FUNCTION "LOWERCASE" : String[254]   // FC273, SCL
TITLE = LOWERCASE
{ S7_Optimized_Access := 'FALSE' }
AUTHOR : hugo
FAMILY : STRINGS
NAME : LOWCASE
VERSION : 1.3
// lowercase returns str while all letters A..Z and Ä.Ö,Ü are converted to lowercase.
//  
// uses: SETUP [DB1]
//       TO_LOWER [FC282]
   VAR_INPUT
      str : String[254];
      _str AT str : Struct
         length : Byte;
         act_length : Byte;
         str : Array[1..254] of Byte;
      END_STRUCT;
   END_VAR
   VAR_TEMP
      tLOWERCASE : String[254];
      _LOWERCASE AT tLOWERCASE : Struct
         length : Byte;
         act_length : Byte;
         str : Array[1..254] of Byte;
      END_STRUCT;
      PT : Int;   // PT : POINTER TO BYTE;
      pos : Int;
      l : Int;
   END_VAR
BEGIN


   #PT := 1;                                    //ADR(LOWERCASE);
   #tLOWERCASE := #str;
   #l := BYTE_TO_INT(#_LOWERCASE.act_length);    //LEN(str);
   FOR #pos := 1 TO #l DO
       #_LOWERCASE.str[#PT] := "TO_LOWER"(#_LOWERCASE.str[#PT]);
       #PT := #PT + 1;
   END_FOR;

   #LOWERCASE := #tLOWERCASE;

   (* revision histroy
   hm  6. oct. 2006    rev 1.0
       original release

   hm  4. feb. 2008    rev 1.1
       improved performance
       added Ä.Ö,Ü

   hm  6. mar. 2008    rev 1.2
       added support for exteded Ascii

   hm  29. mar. 2008   rev 1.3
       changed STRING to STRING(STRING_LENGTH)
   *)
END_FUNCTION

FUNCTION "MIRROR" : String[254]   // FC274, SCL
TITLE = MIRROR
{ S7_Optimized_Access := 'FALSE' }
AUTHOR : hugo
FAMILY : STRINGS
NAME : MIRROR
VERSION : 1.1
// this function reverses an input string.
   VAR_INPUT
      str : String[254];
      _str AT str : Struct
         length : Byte;
         act_length : Byte;
         str : Array[1..254] of Byte;
      END_STRUCT;
   END_VAR
   VAR_TEMP
      tmirror : String[254];
      _mirror AT tmirror : Struct
         length : Byte;
         act_length : Byte;
         str : Array[1..254] of Byte;
      END_STRUCT;
      pi : Int;   // pi : POINTER TO ARRAY[1..255] OF BYTE;
      po : Int;   // po : POINTER TO BYTE;
      lx : Int;
      i : Int;
   END_VAR
BEGIN


   #tmirror := #str;

   #pi := 1;    //ADR(str);
   #po := 1;    //ADR(mirror);
   #lx := BYTE_TO_INT(#_str.act_length); //LEN(str);
   FOR #i := #lx TO 1 BY - 1 DO
       #_mirror.str[#po] := #_str.str[#i];
       #po := #po + 1;
   END_FOR;
   (* close output string *)
   //po^:= 0;
   #MIRROR:= #tmirror;


   (* revision histroy
   hm  4. feb. 2008    rev 1.0
       original release

   hm  29. mar. 2008   rev 1.1
       changed STRING to STRING(STRING_LENGTH)
   *)
END_FUNCTION

FUNCTION "MONTH_TO_STRING" : String[254]   // FC275, SCL
TITLE = MONTH_TO_STRING
{ S7_Optimized_Access := 'FALSE' }
AUTHOR : hugo
FAMILY : STRINGS
NAME : MONTHSTR
VERSION : 1.1
// MONTH_TO_STRING converts an Integer 1..12 into a String with the Names of the corresponding Month.
// the decoding is according to the language setup in global vars
// 
// uses: LANGUAGE [DB4]
   VAR_INPUT
      MTH : Int;
      LANG : Int;
      LX : Int;
   END_VAR
   VAR_TEMP
      ly : Int;
   END_VAR
BEGIN


   #MONTH_TO_STRING := ' ';

   IF #LANG = 0 THEN #ly := "LANGUAGE".DEFAULT; ELSE #ly := MIN(IN1:=#LANG, IN2:="LANGUAGE".LMAX); END_IF;
   IF #MTH < 1 OR #MTH > 12 THEN
       RETURN;
   ELSIF #LX = 0 THEN
       #MONTH_TO_STRING := "LANGUAGE".MONTHS[#ly, #MTH];
   ELSIF #LX = 3 THEN
       #MONTH_TO_STRING := "LANGUAGE".MONTHS3[#ly, #MTH];
   END_IF;


   (* revisison history

   hm  21. sep. 2008   rev 1.0
       original version

   hm  19. oct. 2008   rev 1.1
       changed language setup constants
   *)
END_FUNCTION

FUNCTION "OCT_TO_BYTE" : Byte   // FC276, SCL
TITLE = OCT_TO_BYTE
{ S7_Optimized_Access := 'FALSE' }
AUTHOR : hugo
FAMILY : STRINGS
NAME : OCT2BY
VERSION : 1.1
// OCT_TO_BYTE converts a octagonal string into a byte.
   VAR_INPUT
      OCT : String[254];
      _OCT AT OCT : Struct
         length : Byte;
         act_length : Byte;
         str : Array[1..10] of Byte;
      END_STRUCT;
   END_VAR
   VAR_TEMP
      pt : Int;   // pt : POINTER TO BYTE;
      i : Int;
      X : Byte;
      stop : Int;
   END_VAR
BEGIN


   #pt := 1;    //ADR(oct);
   #stop := BYTE_TO_INT(#_OCT.act_length);    //LEN(oct);
   FOR #i := 1 TO #stop DO
       (* read the first character and subtract 48 to get value in decimal 0 = 48 *)
       #X := #_OCT.str[#pt];
       (* calculate the value of the digit *)
       IF BYTE_TO_INT(#X) > 47 AND BYTE_TO_INT(#X) < 56 THEN
           #OCT_TO_BYTE := INT_TO_BYTE(BYTE_TO_INT(SHL(IN:=#OCT_TO_BYTE,N:=3)) + BYTE_TO_INT(#X) - 48);
       END_IF;
       #pt := #pt + 1;
   END_FOR;



   (* revision histroy
   hm  18. jun. 2008   rev 1.0
       original release

   hm  20. sep. 2008   rev 1.1
       changed length of input string from 20 to 10

   *)
END_FUNCTION

FUNCTION "OCT_TO_DWORD" : DWord   // FC277, SCL
TITLE = OCT_TO_DWORD
{ S7_Optimized_Access := 'FALSE' }
AUTHOR : hugo
FAMILY : STRINGS
NAME : OCT2DW
VERSION : 1.0
// OCT_TO_DWORD converts a octagonal string into a dword.
   VAR_INPUT
      OCT : String[254];
      _OCT AT OCT : Struct
         length : Byte;
         act_length : Byte;
         str : Array[1..20] of Byte;
      END_STRUCT;
   END_VAR
   VAR_TEMP
      pt : Int;   // pt : POINTER TO BYTE;
      i : Int;
      X : Byte;
      stop : Int;
   END_VAR
BEGIN


   #pt := 1;    //ADR(oct);
   #stop := BYTE_TO_INT(#_OCT.act_length);   //LEN(oct);
   FOR #i := 1 TO #stop DO
       (* read the first character and subtract 48 to get value in decimal 0 = 48 *)
       #X := #_OCT.str[#pt];
       (* calculate the value of the digit *)
       IF BYTE_TO_INT(#X) > 47 AND BYTE_TO_INT(#X) < 56 THEN
           #OCT_TO_DWORD := DINT_TO_DWORD(DWORD_TO_DINT(SHL(IN:=#OCT_TO_DWORD,N:=3)) + BYTE_TO_INT(#X) - 48);
       END_IF;
       #pt := #pt + 1;
   END_FOR;




   (* revision histroy
   hm  18. jun. 2008   rev 1.0
       original release


   *)
END_FUNCTION

FUNCTION "REAL_TO_STRF" : String[254]   // FC278, SCL
TITLE = REAL_TO_STRF
{ S7_Optimized_Access := 'FALSE' }
AUTHOR : oscat
FAMILY : STRINGS
NAME : REALSTR
VERSION : 1.7
// Real_to_strF converts a Real to a fixed length String.
// the string will be filles with zeroes to achieve the fixed length after the dot.
// 
// uses: DI_STRNG [FC5]
//       CONCAT [FC2]
//       EXP10 [FC77]
//       DELETE [FC4]
//       INSERT [FC17]
   VAR_INPUT
      IN : Real;
      N : Int;
   END_VAR
   VAR_TEMP
      tN : Int;
      O : Real;
      i : Int;
      str : String[20];
      _str AT str : Struct
         length : Byte;
         act_length : Byte;
         str : Array[1..20] of Byte;
      END_STRUCT;
      tStr : String[20];
   END_VAR
BEGIN


   (* Initialisierung der temporären Strings *)
   #str := '';
   #tStr := '';
   (* round the input to N digits and convert to string *)
   (* LIMIT N to 0 .. 7 *)
   #tN := LIMIT(MN:=0,IN:=#N,MX:=7);
   (* round the input to N digits and convert to string *)
   #O := ABS(#IN) * "EXP10"(#tN);
   #str := S_CONV(REAL_TO_DINT(#O));
   (* Vorzeichen löschen *)
   #tStr := DELETE(IN:=#str, L:=1, P:=1); 
   #str BLKMOV #tStr;
   (* add zeroes in front to make sure sting is at least 8 digits long *)
   FOR #i := BYTE_TO_INT(#_str.act_length) TO #tN DO 
       #tStr := CONCAT(IN1:='0', IN2:=#str);
       #str BLKMOV #tStr; 
   END_FOR;
   (* add a dot if n > 0 *)
   IF #IN <> 0 THEN 
       #tStr := INSERT(IN1:=#str, IN2:='.', P:=BYTE_TO_INT(#_str.act_length) - #tN); 
   END_IF;
   #str BLKMOV #tStr;
   (* add a minus sign if in is negative *)
   IF #IN < 0 THEN 
       #str := CONCAT(IN1:='-', IN2:=#tStr); 
   END_IF;

   #REAL_TO_STRF := #str;


   (* revision history
   hm  26 jan 2007 rev 1.0
       original version

   hm  20. nov. 2007   rev 1.1
       when N=0 ther will be no dot at the end of the string.

   hm  15. dec. 2007   rev 1.2
       changed code for better performance

   hm  4. mar. 2008    rev 1.3
       result is now rounded instead of trunc

   hm  20. mar. 2008   rev 1.4
       changed trunc to real_to_dint because trunc was generating wrong values on wago 842

   hm  29. mar. 2008   rev 1.5
       changed STRING to STRING(20)

   hm  4. apr. 2008    rev 1.6
       added variable O to avoid an error uner CoDeSys SP PLCWinNT V2.4

   hm  27. feb. 2009   rev 1.7
       added a missing zero for IN < 1

   *)
END_FUNCTION

FUNCTION "REPLACE_ALL" : String[254]   // FC279, SCL
TITLE = REPLACE_ALL
{ S7_Optimized_Access := 'FALSE' }
AUTHOR : hugo
FAMILY : STRINGS
NAME : REPLALL
VERSION : 1.1
// the function findP searches a string str for the occurence of src beginning at the position pos.
// 
// uses: LEN [FC21]
//       FINDP [FC248]
//       EQ_STRNG [FC10] 
//       MID [FC26] 
//       REPLACE [FC31]
   VAR_INPUT
      str : String[254];
      src : String[254];
      rep : String[254];
   END_VAR
   VAR_TEMP
      tstr : String[254];
      tsrc : String[254];
      trep : String[254];
      tREPLACE_ALL : String[254];
      pos : Int;
      lp : Int;
      lx : Int;
   END_VAR
BEGIN


   #tstr := #str;
   #tsrc := #src;
   #trep := #rep;

   #tREPLACE_ALL := #str;
   #lx := LEN(#tsrc);
   #lp := LEN(#trep);
   #pos := "FINDP"(str:=#tREPLACE_ALL,src:=#tsrc,pos:=1);
   WHILE #pos > 0 DO
       #tREPLACE_ALL := REPLACE(IN1:=#tREPLACE_ALL,IN2:=#trep,L:=#lx,P:=#pos);
       #pos := "FINDP"(str:=#tREPLACE_ALL,src:=#tsrc,pos:=#pos + #lp);
   END_WHILE;

   #REPLACE_ALL := #tREPLACE_ALL;

   (* revision histroy
   hm  4. feb. 2008    rev 1.0
       original release

   hm  29. mar. 2008   rev 1.1
       changed STRING to STRING(STRING_LENGTH)
   *)
END_FUNCTION

FUNCTION "REPLACE_CHARS" : String[254]   // FC280, SCL
TITLE = REPLACE_CHARS
{ S7_Optimized_Access := 'FALSE' }
AUTHOR : hugo
FAMILY : STRINGS
NAME : REPLCHR
VERSION : 1.0
// REPLACE_CHARS erstezt alle character die im string src aufgeführt sind mit dem an der selben stelle im string rep gelisteten character.
// 
// uses: TEMP [DB7]
//       LEN [FC21]
//       LEFT [FC20]
//       MID [FC26]
//       FIND [FC11]
//       REPLACE [FC31]
   VAR_INPUT
      STR : String[254];
      SRC : String[254];
      REP : String[254];
   END_VAR
   VAR_TEMP
      "a" : Int;
      "b" : Int;
      c : String[1];
      stp : Int;
   END_VAR
BEGIN


   "TEMP".STR1 := #STR;
   "TEMP".STR2 := #SRC;
   "TEMP".STR3 := #REP;

   "TEMP".TEMP := #STR;
   (* make sure rep and src are of same length and length is > 0 *)
   #"a" := LEN("TEMP".STR1);
   #"b" := LEN("TEMP".STR3);
   IF #"a" < #"b" THEN
       "TEMP".STR3 := LEFT(IN:="TEMP".STR3, L:=#"a");
   ELSIF #"b" < #"a" THEN
       "TEMP".STR2 := LEFT(IN:="TEMP".STR2, L:=#"b");
   END_IF;

   (* search the string and replace if necessary *)
   #stp := LEN("TEMP".STR1);
   FOR #"a" := 1 TO #stp DO
       #c := MID(IN:="TEMP".TEMP, L:=1, P:=#"a");
       #"b" := FIND(IN1:="TEMP".STR2, IN2:=#c);
       IF #"b" > 0 THEN
           "TEMP".TEMP := REPLACE(IN1:="TEMP".TEMP, IN2:=MID(IN:="TEMP".STR3, L:=1, P:=#"b"), L:=1, P:=#"a");
       END_IF;
   END_FOR;

   #REPLACE_CHARS := "TEMP".TEMP;

   (* revision history
   hm      14. may. 2008   rev 1.0
       original version

   *)
END_FUNCTION

FUNCTION "REPLACE_UML" : String[254]   // FC281, SCL
TITLE = REPLACE_UML
{ S7_Optimized_Access := 'FALSE' }
AUTHOR : kurt
FAMILY : STRINGS
NAME : REPLUML
VERSION : 1.1
// REPLACE_UML replaces all occurences of Ä,Ö,Ü and ä,ö,ü,ß with Ae, ae, Oe, oe, Ue, ue and ss.
// 
// uses: TO_UML [FC283]
//       CHR_TO_STRING [FC227]
   VAR_INPUT
      str : String[254];
      _str AT str : Struct
         length : Byte;
         act_length : Byte;
         str : Array[1..254] of Byte;
      END_STRUCT;
   END_VAR
   VAR_TEMP
      tREPLACE_UML : String[254];
      _REPLACE_UML AT tREPLACE_UML : Struct
         length : Byte;
         act_length : Byte;
         str : Array[1..254] of Byte;
      END_STRUCT;
      l : Int;
      pt : Int;   // pt : POINTER TO BYTE;
      pto : Int;   // pto : POINTER TO BYTE;
      ptm : Int;   // ptm : POINTER TO BYTE;
      pt1 : Int;   // pt1, pt2 : POINTER TO BYTE;
      pt2 : Int;   // pt1, pt2 : POINTER TO BYTE;
      su : String[2];
      _su AT su : Struct
         length : Byte;
         act_length : Byte;
         str : Array[1..2] of Byte;
      END_STRUCT;
      pos : Int;
   END_VAR
BEGIN


   #tREPLACE_UML := #str;

   #pt := 1;    //ADR(str);
   #pto := 1;   //ADR(REPLACE_UML);
   #ptm := #pto; // + INT_TO_DWORD(string_length);
   #pt1 := 1;   //ADR(su);
   #pt2 := #pt1 + 1;
   #l := BYTE_TO_INT(#_str.act_length);   //LEN(str);
   WHILE #pos < #l AND #pos < BYTE_TO_INT(#_str.act_length) DO
       IF BYTE_TO_INT(#_str.str[#pt]) < 127 THEN
           (* no uml character simlply copy the character*)
           #_REPLACE_UML.str[#pto] := #_str.str[#pt];
       ELSE
           (* convert the uml character *)
           #su := "TO_UML"(#_str.str[#pt]);
           (* we must make sure pointer are not out of range *)
           #_REPLACE_UML.str[#pto] := #_su.str[#pt1];
           IF #pto < #ptm THEN
               #pto := #pto + 1;
               #_REPLACE_UML.str[#pto] := #_su.str[#pt2];
           END_IF;
       END_IF;
       (* increment pointers *)
       #pt := #pt + 1;
       #pto := #pto + 1;
       #pos := #pos + 1;
   END_WHILE;

   (* properly close the output string *)
   //pto^ := 0;
   #REPLACE_UML := #tREPLACE_UML;

   (* revision history
   hm  29. feb 2008    rev 1.0
       original version

   hm  29. mar. 2008   rev 1.1
       changed STRING to STRING(STRING_LENGTH)
       new code to avoid pointer out of range
       use new function to_uml
   *)
END_FUNCTION

FUNCTION "TO_LOWER" : Byte   // FC282, SCL
TITLE = TO_LOWER
{ S7_Optimized_Access := 'FALSE' }
AUTHOR : hugo
FAMILY : STRINGS
NAME : TO_LOWER
VERSION : 1.2
// to_lower converts a character from uppercase to lowercase
// 
// uses: SETUP [DB1]
   VAR_INPUT
      IN : Byte;
   END_VAR
BEGIN


   IF BYTE_TO_INT(#IN) > 64 AND BYTE_TO_INT(#IN) < 91 THEN
      #TO_LOWER := #IN OR 16#20;
   ELSIF (BYTE_TO_INT(#IN) > 191 AND BYTE_TO_INT(#IN) < 223) AND BYTE_TO_INT(#IN) <> 215 AND "SETUP".EXTENDED_ASCII THEN
      #TO_LOWER := #IN OR 16#20;
   ELSE
      #TO_LOWER := #IN;
   END_IF;


   (* revision history
   hm  6. mar. 2008    rev 1.0
       original version

   hm  19. oct. 2008   rev 1.1
       changed setup constants

   ks  25. oct. 2008   rev 1.2
       optimized code
   *)
END_FUNCTION

FUNCTION "TO_UML" : String[254]   // FC283, SCL
TITLE = TO_UML
{ S7_Optimized_Access := 'FALSE' }
AUTHOR : hugo
FAMILY : STRINGS
NAME : TO_UML
VERSION : 1.1
// to_uml converts a character above 127 to a two digit character below 127.
// the character Ä is converted to Ae
// 
// uses: CHR_TO_STRING [FC227]
   VAR_INPUT
      IN : Byte;
   END_VAR
   VAR_TEMP
      tTO_UML : String[2];
   END_VAR
BEGIN


   CASE BYTE_TO_INT(#IN) OF
       196:    (* Ä *)
           #tTO_UML := 'Ae';
       214:    (* Ö *)
           #tTO_UML := 'Oe';
       220:    (* Ü *)
           #tTO_UML := 'Ue';
       223:    (* ß *)
           #tTO_UML := 'ss';
       228:    (* ä *)
           #tTO_UML := 'ae';
       246:    (* ö *)
           #tTO_UML := 'oe';
       252:    (* ü *)
           #tTO_UML := 'ue';
   ELSE
       #tTO_UML := "CHR_TO_STRING"(#IN);
   END_CASE;

   #TO_UML := #tTO_UML;


   (* revision history
   hm  29. mar. 2008   rev 1.0
       original version

   hm  17. dec. 2008   rev 1.1
       changes name of function chr to chr_to_string

   *)
END_FUNCTION

FUNCTION "TO_UPPER" : Byte   // FC284, SCL
TITLE = TO_UPPER
{ S7_Optimized_Access := 'FALSE' }
AUTHOR : hugo
FAMILY : STRINGS
NAME : TO_UPPER
VERSION : 1.3
// to_upper converts a character from lowercase to uppercase
// 
// uses: SETUP [DB1]
   VAR_INPUT
      IN : Byte;
   END_VAR
BEGIN


   IF BYTE_TO_INT(#IN) > 96 AND BYTE_TO_INT(#IN) < 123 THEN
      #TO_UPPER := #IN AND 16#DF;
   ELSIF BYTE_TO_INT(#IN) > 223 AND BYTE_TO_INT(#IN) <> 247 AND BYTE_TO_INT(#IN) <> 255 AND "SETUP".EXTENDED_ASCII THEN
      #TO_UPPER := #IN AND 16#DF;
   ELSE
      #TO_UPPER := #IN;
   END_IF;


   (* revision history
   hm  6. mar. 2008    rev 1.0
       original version

   hm  19. oct. 2008   rev 1.1
       changed setup constants

   ks  25. oct. 2008   rev 1.2
       optimized code

   hm 16. jan 2009 rev 1.3
       corrected an error in module

   *)
END_FUNCTION

FUNCTION "TRIM" : String[254]   // FC285, SCL
TITLE = TRIM
{ S7_Optimized_Access := 'FALSE' }
AUTHOR : hugo
FAMILY : STRINGS
NAME : TRIM
VERSION : 1.2
// the function deletes all blanks within a string.
// 
// uses: FIND [FC11]
//       REPLACE [FC31]
   VAR_INPUT
      str : String[254];
   END_VAR
   VAR_TEMP
      tstr : String[254];
      pos : Int;
   END_VAR
BEGIN


   #tstr := #str;

   REPEAT
       #pos := FIND(IN1:=#tstr,IN2:=' ');
       IF #pos > 0 THEN #tstr := REPLACE(IN1:=#tstr,IN2:='',L:=1,P:=#pos); END_IF;
   UNTIL #pos = 0   END_REPEAT;

   #TRIM := #tstr;


   (* revision histroy
   hm  6.10.2006       rev 1.0
       original release

   hm  20. mar. 2008   rev 1.1
       avoid to call replace with pos = 0 because some systems will produce an error

   hm  29. mar. 2008   rev 1.2
       changed STRING to STRING(STRING_LENGTH)
   *)
END_FUNCTION

FUNCTION "TRIM1" : String[254]   // FC286, SCL
TITLE = TRIM1
{ S7_Optimized_Access := 'FALSE' }
AUTHOR : hugo
FAMILY : STRINGS
NAME : TRIM1
VERSION : 1.2
// the function replaces all multiple blanks within a string by only one blank.
// leading and ending blanks will be deleted
// 
// uses: EQ_STRNG [FC10]
//       FIND [FC11]
//       REPLACE [FC31]
//       LEFT [FC20]
//       DELETE [FC4]
//       RIGHT [FC32]
//       LEN [FC21]
   VAR_INPUT
      str : String[254];
   END_VAR
   VAR_TEMP
      tstr : String[254];
      pos : Int;
   END_VAR
BEGIN


   #tstr := #str;

   REPEAT
       #pos := FIND(IN1:=#tstr,IN2:='  ');
       IF #pos > 0 THEN #tstr := REPLACE(IN1:=#tstr,IN2:=' ',L:=2,P:=#pos); END_IF;
   UNTIL #pos = 0   END_REPEAT;
   (* beginning and ending blanks need to be stripped off *)
   IF LEFT(IN:=#tstr,L:=1) S_COMP ' ' THEN #tstr := DELETE(IN:=#tstr,L:=1,P:=1); END_IF;
   IF RIGHT(IN:=#tstr,L:=1) S_COMP ' ' THEN #tstr := DELETE(IN:=#tstr,L:=1,P:=LEN(#tstr)); END_IF;

   #TRIM1 := #tstr;

   (* revision histroy
   hm  4. feb. 2008    rev 1.0
       original release

   hm  20. mar. 2008   rev 1.1
       avoid to call replace with pos = 0 because some systems will produce an error

   hm  29. mar. 2008   rev 1.2
       changed STRING to STRING(STRING_LENGTH)
   *)
END_FUNCTION

FUNCTION "TRIME" : String[254]   // FC287, SCL
TITLE = TRIME
{ S7_Optimized_Access := 'FALSE' }
AUTHOR : hugo
FAMILY : STRINGS
NAME : TRIME
VERSION : 1.0
// this function deletes all leading and ending blanks of a string.
//  
// uses: TEMP [DB7]
//       EQ_STRNG [FC10]
//       LEFT [FC20]
//       DELETE [FC4]
//       RIGHT [FC32]
//       LEN [FC21]
   VAR_INPUT
      str : String[254];
   END_VAR
BEGIN


   "TEMP".STR1 := #str;
   (* beginning blanks need to be stripped off *)
   WHILE LEFT(IN:="TEMP".STR1,L:=1) S_COMP ' ' DO
       "TEMP".STR1 := DELETE(IN:="TEMP".STR1,L:=1,P:=1);
   END_WHILE;

   (* ending blanks need to be stripped off *)
   WHILE RIGHT(IN:="TEMP".STR1,L:=1) S_COMP ' ' DO
       "TEMP".STR1 := DELETE(IN:="TEMP".STR1,L:=1,P:=LEN("TEMP".STR1));
   END_WHILE;

   #TRIME := "TEMP".STR1;

   (* revision histroy
   hm  28. mar. 2008   rev 1.0
       original release

   *)
END_FUNCTION

FUNCTION "UPPERCASE" : String[254]   // FC288, SCL
TITLE = UPPERCASE
{ S7_Optimized_Access := 'FALSE' }
AUTHOR : hugo
FAMILY : STRINGS
NAME : UPCASE
VERSION : 1.3
// uppercase returns str while all letters a..z and ä,ö,ü are converted to uppercase
// 
// uses: SETUP [DB1]
//       TO_UPPER [FC284]
   VAR_INPUT
      str : String[254];
   END_VAR
   VAR_TEMP
      tUPPERCASE : String[254];
      _UPPERCASE AT tUPPERCASE : Struct
         length : Byte;
         act_length : Byte;
         str : Array[1..254] of Byte;
      END_STRUCT;
      PT : Int;   // PT : POINTER TO BYTE;
      pos : Int;
      l : Int;
   END_VAR
BEGIN


   #PT := 1;
   #tUPPERCASE := #str;
   #l := BYTE_TO_INT(#_UPPERCASE.act_length);
   FOR #pos := 1 TO #l DO
       #_UPPERCASE.str[#PT] := "TO_UPPER"(#_UPPERCASE.str[#PT]);
       #PT := #PT + 1;
   END_FOR;

   #UPPERCASE := #tUPPERCASE;

   (* revision histroy
   hm  6. oct. 2006    rev 1.0
       original release

   hm  4. feb. 2008    rev 1.1
       improved performance
       added Ä,Ö,Ü

   hm  6. mar. 2008    rev 1.2
       added support for exteded Ascii

   hm  29. mar. 2008   rev 1.3
       changed STRING to STRING(STRING_LENGTH)
   *)
END_FUNCTION

FUNCTION "WEEKDAY_TO_STRING" : String[254]   // FC289, SCL
TITLE = WEEKDAY_TO_STRING
{ S7_Optimized_Access := 'FALSE' }
AUTHOR : hugo
FAMILY : STRINGS
NAME : WDSTR
VERSION : 1.1
// WEEKDAY_TO_STRING converts an Integer 1..7 into a String with the Names of the corresponding weekday.
// the decoding is according to the language setup in global vars
// 
// uses: LANGUAGE [DB4]
   VAR_INPUT
      WDAY : Int;
      LANG : Int;
      LX : Int;
   END_VAR
   VAR_TEMP
      ly : Int;
   END_VAR
BEGIN


   IF #LANG = 0 THEN #ly := "LANGUAGE".DEFAULT; ELSE #ly := MIN(IN1:=#LANG, IN2:="LANGUAGE".LMAX); END_IF;
   IF #WDAY < 1 OR #WDAY > 7 THEN
       RETURN;
   ELSIF #LX = 0 THEN
       #WEEKDAY_TO_STRING := "LANGUAGE".WEEKDAYS[#ly, #WDAY];
   ELSIF #LX = 2 THEN
       #WEEKDAY_TO_STRING := "LANGUAGE".WEEKDAYS2[#ly, #WDAY];
   END_IF;


   (* revisison history

   hm  21. sep. 2008   rev 1.0
       original version

   hm  19. oct. 2008   rev 1.1
       changed language setup constants
   *)
END_FUNCTION

FUNCTION "FSTRING_TO_DT" : Date_And_Time   // FC403, SCL
TITLE = FSTRING_TO_DT
{ S7_Optimized_Access := 'FALSE' }
AUTHOR : hugo
FAMILY : STRINGS
NAME : FSTR2DT
VERSION : 1.0
// FSTRING_TO_DT converts Formatted String into a DT value.
// 
// uses: TEMP [DB7]
//       SETUP [DB1]
//       LANGUAGE [DB4]
//       STRNG_I [FC38]
//       EQ_STRNG [FC10]
//       TRIM [FC285]
//       FIND [FC11] 
//       REPLACE [FC31] 
//       CAPITALIZE [FC224]
//       TO_UPPER [FC284] 
//       LOWERCASE [FC273]
//       TO_LOWER [FC282] 
//       NE_STRNG [FC29]
//       LEFT [FC20]
//       DELETE [FC4]
//       MID [FC26]
//       SET_DT [FC214]
   VAR_INPUT
      SDT : String[254];
      FMT : String[254];
   END_VAR
   VAR_TEMP
      tFSTRING_TO_DT : Date_And_Time;
      c : String[1];
      tmp : String[20];
      end : Int;
      dy : Int;
      dm : Int;
      dd : Int;
      th : Int;
      tm : Int;
      ts : Int;
   END_VAR
BEGIN


   "TEMP".STR1 := #SDT;
   "TEMP".STR2 := #FMT;
   #tmp := '';

   (* scan input string *)
   WHILE "TEMP".STR2 <> '' DO
       #c := LEFT(IN:="TEMP".STR2,L:=1);
       IF #c = '*' THEN //ignore
           (* skip ignore characters *)
           "TEMP".STR2 := DELETE(IN:="TEMP".STR2,L:=1,P:=1);
           "TEMP".STR1 := DELETE(IN:="TEMP".STR1,L:=1,P:=1);
       ELSIF #c = '#' THEN //fchar
           (* format chracter found skip format char and read identifier *)
           (* store format identifier in c and skip to next char in fmt *)
           #c := MID(IN:="TEMP".STR2,L:=1,P:=2);
           "TEMP".STR2 := DELETE(IN:="TEMP".STR2,L:=2,P:=1);
           (* extract the substring until the end of sdt or to next char of fmt *)
           IF "TEMP".STR2 = '' THEN
               #tmp := "TEMP".STR1;
           ELSE
               (* serach for end of substring *)
               #end := FIND(IN1:="TEMP".STR1, IN2:=LEFT(IN:="TEMP".STR2, L:=1))-1;
               #tmp := LEFT(IN:="TEMP".STR1, L:=#end);
               "TEMP".STR1 := DELETE(IN:="TEMP".STR1, L:=#end, P:=1);
           END_IF;
           (* extract information from substring *)
           IF #c = 'Y' THEN
               #dy := S_CONV(#tmp);
               IF #dy < 100 THEN #dy := #dy + 2000; END_IF;
           ELSIF #c = 'M' THEN
               #dm := S_CONV(#tmp);
           ELSIF #c = 'N' THEN
               #dm := "FSTRING_TO_MONTH"(MTH:=#tmp,LANG:=0);
           ELSIF #c = 'D' THEN
               #dd := S_CONV(#tmp);
           ELSIF #c = 'h' THEN
               #th := S_CONV(#tmp);
           ELSIF #c = 'm' THEN
               #tm := S_CONV(#tmp);
           ELSIF #c = 's' THEN
               #ts := S_CONV(#tmp);
           END_IF;
       ELSIF #c = LEFT(IN:="TEMP".STR1,L:=1) THEN
           (* skip matching characters *)
           "TEMP".STR2 := DELETE(IN:="TEMP".STR2,L:=1,P:=1);
           "TEMP".STR1 := DELETE(IN:="TEMP".STR1,L:=1,P:=1);
       ELSE
           RETURN;
       END_IF;
   END_WHILE;

   #tFSTRING_TO_DT := "SET_DT"(year:=#dy,month:=#dm,day:=#dd,hour:=#th,minute:=#tm,second:=#ts);
   #FSTRING_TO_DT := #tFSTRING_TO_DT;

   (* revision histroy
   hm  24. sep. 2008   rev 1.0
       original release


   *)
END_FUNCTION

FUNCTION "DATE_DINT" : DInt   // FC405, SCL
TITLE = DATE_DINT
{ S7_Optimized_Access := 'FALSE' }
AUTHOR : dalbi
FAMILY : xS7
NAME : D_DINT
VERSION : 1.0
// convert S7 DATE to IEC-DATE
   VAR_INPUT
      D : Date;
   END_VAR
BEGIN


   (* 1.1.1990 00:00:00 = 631152000 *)
   #DATE_DINT := T_CONV(#D) * 86400 + 631152000;
END_FUNCTION

FUNCTION "COUNT_SUBSTRING" : Int   // FC433, SCL
TITLE = COUNT_SUBSTRING
{ S7_Optimized_Access := 'FALSE' }
AUTHOR : kurt
FAMILY : STRINGS
NAME : CTSUBSTR
VERSION : 1.0
// count_substring returns the number of occurences of a substring in a string
// 
// uses: LEN (FC21)
//       FIND (FC11)
//       REPLACE (FC31)
   VAR_INPUT
      SEARCH : String[254];
      STR : String[254];
   END_VAR
   VAR_TEMP
      pos : Int;
      size : Int;
   END_VAR
BEGIN


   "TEMP".STR1 := #SEARCH;
   "TEMP".STR2 := #STR;

   #COUNT_SUBSTRING := 0;
   #size := LEN("TEMP".STR1);
   REPEAT
      #pos := FIND(IN1:="TEMP".STR2,IN2:="TEMP".STR1);
      IF #pos > 0 THEN
         "TEMP".STR2 := REPLACE(IN1:="TEMP".STR2,IN2:='',L:=#size,P:=#pos);
         #COUNT_SUBSTRING := #COUNT_SUBSTRING + 1;
      END_IF;
   UNTIL #pos = 0
   END_REPEAT;


   (* revision history
   ks  20. jan. 2011 rev 1.0
     original version

   *)
END_FUNCTION

// ===== PLC "Time and Date"  Unspecific CPU S7 300 =====

VAR_GLOBAL CONSTANT   // PLC tag table "STEP7 classic symbols"
   "MTH_OFS1" : Int := 0;
   "MTH_OFS2" : Int := 31;
   "MTH_OFS3" : Int := 59;
   "MTH_OFS4" : Int := 90;
   "MTH_OFS5" : Int := 120;
   "MTH_OFS6" : Int := 151;
   "MTH_OFS7" : Int := 181;
   "MTH_OFS8" : Int := 212;
   "MTH_OFS9" : Int := 243;
   "MTH_OFS10" : Int := 273;
   "MTH_OFS11" : Int := 304;
   "MTH_OFS12" : Int := 334;
   "PI2" : Real := 6.283185307179586476;   // PI * 2
   "PI" : Real := 3.14159265358979323846264338327950288;   // Kreiszahl PI
   "PI2_FB31" : Real := 6.28318530717958647692528676655900576;   // MigChange: PI2 OriginalComment: PI * 2
   "debug" : Bool := FALSE;
   "N" : Int := 0;
   "offset" : Int := 0;
   "offset_1" : DWord := 0;
END_VAR

TYPE "CALENDAR"
VERSION : 0.0
   STRUCT
      UTC : Date_And_Time;   // world time UTC
      LDT : Date_And_Time;   // local time
      LDATE : Date;   // local date
      LTOD : Time_Of_Day;   // local time of day
      YEAR : Int;   // year of LDATE
      MONTH : Int;   // month of LDATE
      DAY : Int;   // day of LDATE
      WEEKDAY : Int;   // weekday of LDATE
      OFFSET : Int;   // Time Zone Offset for Local time in minutes
      DST_EN : Bool;   // daylight savings time enable
      DST_ON : Bool;   // true when daylight savings time os on
      _NAME : String[5];   // name of time zone
      LANGUAGE : Int;   // location number pls see location setup
      LONGITUDE : Real;   // longitude of current location
      LATITUDE : Real;   // latitude of current location
      SUN_RISE : Time_Of_Day;   // sun_rise for current location
      SUN_SET : Time_Of_Day;   // sun_set for current location
      SUN_MIDDAY : Time_Of_Day;   // worldtime when sun stands at south position
      SUN_HEIGTH : Real;   // suns heigth at midday, south position
      SUN_HOR : Real;   // sun angle horizontal 0 = north in degrees
      SUN_VER : Real;   // sun angle vertical above horizon in degrees
      NIGHT : Bool;   // true between sun_set and sun_rise
      HOLIDAY : Bool;   // true when holiday
      HOLY_NAME : String[30];   // name of holiday
      WORK_WEEK : Int;   // current work week
   END_STRUCT;
END_TYPE

TYPE "HOLIDAY_DATA"
VERSION : 0.0
   STRUCT
      _NAME : String[30];
      DAY : Int;
      MONTH : Int;
      USE : Int;
   END_STRUCT;
END_TYPE

TYPE "SDT"
VERSION : 0.0
   STRUCT
      YEAR : Int;
      MONTH : Int;
      DAY : Int;
      WEEKDAY : Int;
      HOUR : Int;
      MINUTE : Int;
      SECOND : Int;
      MS : Int;
   END_STRUCT;
END_TYPE

DATA_BLOCK "LANGUAGE"   // DB4
TITLE = LANGUAGE
{ S7_Optimized_Access := 'FALSE' }
AUTHOR : oscat
FAMILY : CONSTANT
NAME : DBLANG
VERSION : 1.2
   VAR
      DEFAULT : Int := 1;   // 1=english, 2=german, 3=french
      LMAX : Int := 3;
      WEEKDAYS : Array[1..3, 1..7] of String[10];
      WEEKDAYS2 : Array[1..3, 1..7] of String[2];
      MONTHS : Array[1..3, 1..12] of String[10];
      MONTHS3 : Array[1..3, 1..12] of String[3];
      DIRS : Array[1..3, 0..15] of String[3];
   END_VAR
BEGIN
   WEEKDAYS[1,1] := 'Monday';
   WEEKDAYS[1,2] := 'Tuesday';
   WEEKDAYS[1,3] := 'Wednesday';
   WEEKDAYS[1,4] := 'Thursday';
   WEEKDAYS[1,5] := 'Friday';
   WEEKDAYS[1,6] := 'Saturday';
   WEEKDAYS[1,7] := 'Sunday';
   WEEKDAYS[2,1] := 'Montag';
   WEEKDAYS[2,2] := 'Dienstag';
   WEEKDAYS[2,3] := 'Mittwoch';
   WEEKDAYS[2,4] := 'Donnerstag';
   WEEKDAYS[2,5] := 'Freitag';
   WEEKDAYS[2,6] := 'Samstag';
   WEEKDAYS[2,7] := 'Sonntag';
   WEEKDAYS[3,1] := 'Lundi';
   WEEKDAYS[3,2] := 'Mardi';
   WEEKDAYS[3,3] := 'Mercredi';
   WEEKDAYS[3,4] := 'Jeudi';
   WEEKDAYS[3,5] := 'Vendredi';
   WEEKDAYS[3,6] := 'Samedi';
   WEEKDAYS[3,7] := 'Dimanche';
   WEEKDAYS2[1,1] := 'Mo';
   WEEKDAYS2[1,2] := 'Tu';
   WEEKDAYS2[1,3] := 'We';
   WEEKDAYS2[1,4] := 'Th';
   WEEKDAYS2[1,5] := 'Fr';
   WEEKDAYS2[1,6] := 'Sa';
   WEEKDAYS2[1,7] := 'Su';
   WEEKDAYS2[2,1] := 'Mo';
   WEEKDAYS2[2,2] := 'Di';
   WEEKDAYS2[2,3] := 'Mi';
   WEEKDAYS2[2,4] := 'Do';
   WEEKDAYS2[2,5] := 'Fr';
   WEEKDAYS2[2,6] := 'Sa';
   WEEKDAYS2[2,7] := 'So';
   WEEKDAYS2[3,1] := 'Lu';
   WEEKDAYS2[3,2] := 'Ma';
   WEEKDAYS2[3,3] := 'Me';
   WEEKDAYS2[3,4] := 'Je';
   WEEKDAYS2[3,5] := 'Ve';
   WEEKDAYS2[3,6] := 'Sa';
   WEEKDAYS2[3,7] := 'Di';
   MONTHS[1,1] := 'January';
   MONTHS[1,2] := 'February';
   MONTHS[1,3] := 'March';
   MONTHS[1,4] := 'April';
   MONTHS[1,5] := 'May';
   MONTHS[1,6] := 'June';
   MONTHS[1,7] := 'July';
   MONTHS[1,8] := 'August';
   MONTHS[1,9] := 'September';
   MONTHS[1,10] := 'October';
   MONTHS[1,11] := 'November';
   MONTHS[1,12] := 'December';
   MONTHS[2,1] := 'Januar';
   MONTHS[2,2] := 'Februar';
   MONTHS[2,3] := 'März';
   MONTHS[2,4] := 'April';
   MONTHS[2,5] := 'Mai';
   MONTHS[2,6] := 'Juni';
   MONTHS[2,7] := 'Juli';
   MONTHS[2,8] := 'August';
   MONTHS[2,9] := 'September';
   MONTHS[2,10] := 'Oktober';
   MONTHS[2,11] := 'November';
   MONTHS[2,12] := 'Dezember';
   MONTHS[3,1] := 'Janvier';
   MONTHS[3,2] := 'Février';
   MONTHS[3,3] := 'mars';
   MONTHS[3,4] := 'Avril';
   MONTHS[3,5] := 'Mai';
   MONTHS[3,6] := 'Juin';
   MONTHS[3,7] := 'Juillet';
   MONTHS[3,8] := 'Août';
   MONTHS[3,9] := 'Septembre';
   MONTHS[3,10] := 'Octobre';
   MONTHS[3,11] := 'Novembre';
   MONTHS[3,12] := 'Decembre';
   MONTHS3[1,1] := 'Jan';
   MONTHS3[1,2] := 'Feb';
   MONTHS3[1,3] := 'Mar';
   MONTHS3[1,4] := 'Apr';
   MONTHS3[1,5] := 'May';
   MONTHS3[1,6] := 'Jun';
   MONTHS3[1,7] := 'Jul';
   MONTHS3[1,8] := 'Aug';
   MONTHS3[1,9] := 'Sep';
   MONTHS3[1,10] := 'Oct';
   MONTHS3[1,11] := 'Nov';
   MONTHS3[1,12] := 'Dec';
   MONTHS3[2,1] := 'Jan';
   MONTHS3[2,2] := 'Feb';
   MONTHS3[2,3] := 'Mrz';
   MONTHS3[2,4] := 'Apr';
   MONTHS3[2,5] := 'Mai';
   MONTHS3[2,6] := 'Jun';
   MONTHS3[2,7] := 'Jul';
   MONTHS3[2,8] := 'Aug';
   MONTHS3[2,9] := 'Sep';
   MONTHS3[2,10] := 'Okt';
   MONTHS3[2,11] := 'Nov';
   MONTHS3[2,12] := 'Dez';
   MONTHS3[3,1] := 'Jan';
   MONTHS3[3,2] := 'Fev';
   MONTHS3[3,3] := 'Mar';
   MONTHS3[3,4] := 'Avr';
   MONTHS3[3,5] := 'Mai';
   MONTHS3[3,6] := 'Jun';
   MONTHS3[3,7] := 'Jul';
   MONTHS3[3,8] := 'Aou';
   MONTHS3[3,9] := 'Sep';
   MONTHS3[3,10] := 'Oct';
   MONTHS3[3,11] := 'Nov';
   MONTHS3[3,12] := 'Dec';
   DIRS[1,0] := 'N';
   DIRS[1,1] := 'NNE';
   DIRS[1,2] := 'NE';
   DIRS[1,3] := 'ENE';
   DIRS[1,4] := 'E';
   DIRS[1,5] := 'ESE';
   DIRS[1,6] := 'SE';
   DIRS[1,7] := 'SSE';
   DIRS[1,8] := 'S';
   DIRS[1,9] := 'SSW';
   DIRS[1,10] := 'SW';
   DIRS[1,11] := 'WSW';
   DIRS[1,12] := 'W';
   DIRS[1,13] := 'WNW';
   DIRS[1,14] := 'NW';
   DIRS[1,15] := 'NNW';
   DIRS[2,0] := 'N';
   DIRS[2,1] := 'NNO';
   DIRS[2,2] := 'NO';
   DIRS[2,3] := 'ONO';
   DIRS[2,4] := 'O';
   DIRS[2,5] := 'OSO';
   DIRS[2,6] := 'SO';
   DIRS[2,7] := 'SSO';
   DIRS[2,8] := 'S';
   DIRS[2,9] := 'SSW';
   DIRS[2,10] := 'SW';
   DIRS[2,11] := 'WSW';
   DIRS[2,12] := 'W';
   DIRS[2,13] := 'WNW';
   DIRS[2,14] := 'NW';
   DIRS[2,15] := 'NNW';
   DIRS[3,0] := 'N';
   DIRS[3,1] := 'NNO';
   DIRS[3,2] := 'NO';
   DIRS[3,3] := 'ONO';
   DIRS[3,4] := 'O';
   DIRS[3,5] := 'OSO';
   DIRS[3,6] := 'SO';
   DIRS[3,7] := 'SSO';
   DIRS[3,8] := 'S';
   DIRS[3,9] := 'SSW';
   DIRS[3,10] := 'SW';
   DIRS[3,11] := 'WSW';
   DIRS[3,12] := 'W';
   DIRS[3,13] := 'WNW';
   DIRS[3,14] := 'NW';
   DIRS[3,15] := 'NNW';
END_DATA_BLOCK

DATA_BLOCK "LOCATION"   // DB5
TITLE = LOCATION
{ S7_Optimized_Access := 'FALSE' }
AUTHOR : oscat
FAMILY : CONSTANT
NAME : DBLOCA
VERSION : 1.2
   VAR
      DEFAULT : Int := 1;   // 1=germany, 2=austria 3=france 4=belgium-german 5= italien-Südtirol
      LMAX : Int := 5;   // language spoken in the location
      LANGUAGE : Array[1..5] of Int;
   END_VAR
BEGIN
   LANGUAGE[1] := 2;
   LANGUAGE[2] := 2;
   LANGUAGE[3] := 3;
   LANGUAGE[4] := 2;
   LANGUAGE[5] := 2;
END_DATA_BLOCK

DATA_BLOCK "IDB_STIME"   // DB64
{ S7_Optimized_Access := 'FALSE' }
AUTHOR : dalbi
FAMILY : MEASURE
VERSION : 0.0
// stored: InstanceOfName STIME
"STIME"
BEGIN
END_DATA_BLOCK

FUNCTION_BLOCK "CALENDAR_CALC"   // FB26, SCL
TITLE = CALENDAR_CALC
{ S7_Optimized_Access := 'FALSE' }
AUTHOR : oscat
FAMILY : TIDT
NAME : CALCALC
VERSION : 1.6
// calendar_calc liest die weltzeit .UTC aus einer CALENDAR Struktur und berechnet die restlichen Werte der Struktur.
// calendar_calc stellt sicher das die Werte fortlaufend aktualisiert werden und dabei funktionen nur dann aufgerufen werden wenn dies nötig ist.
// calendar_calc will calculate sun position data when SPE = TRUE;
// 
// uses: LOCATION [DB5]
//       HOLIDAY_DATA [UDT9]
//       NE_DT [FC28]
//       SB_DT_DT [FC34]
//       DT_TOD [FC8]
//       UTC_TO_LTIME [FC402]
//       DST [FC183] 
//       YEAR_OF_DATE [FC219]
//       DT_DATE [FC6]
//       DT_DINT [FC400]
//       SET_DT [FC214]
//       DINT_DT [FC399] 
//       D_TOD_DT [FC3]
//       DAY_OF_DATE [FC177]
//       HOUR [FC187]
//       MONTH_OF_DATE [FC202]
//       DAY_OF_YEAR [FC180] 
//       YEAR_BEGIN [FC217]
//       LEAP_OF_DATE [FC193] 
//       LEAP_YEAR [FC194]
//       DAY_OF_MONTH [FC178]
//       DAY_OF_WEEK [FC179]
//       HOLIDAY [FB28]
//       EASTER [FC186] 
//       SET_DATE [FC213]
//       DATE_ADD [FC176] 
//       FLOOR [FC81]
//       SGN [FC106]
//       SUN_TIME [FB32]
//       HOUR_TO_TOD [FC190] 
//       WORK_WEEK [FC216]
//       SUN_POS [FB31]
//       MODR [FC97] 
//       FLOOR2 [FC82]
//       RAD [FC100] 
//       DEG [FC72] 
//       REFRACTION [FC206]
   VAR_INPUT
      SPE : Bool;
      H : Real := -8.333333e-1;
   END_VAR
   VAR_IN_OUT
      XCAL : "CALENDAR";
      HOLIDAYS : Array[0..29] of "HOLIDAY_DATA";
   END_VAR
   VAR
      last : Date_And_Time;
      last_day : DInt;
      holy : "HOLIDAY";
      sun : "SUN_TIME";
      last_hour : Int;
      utod : Time_Of_Day;
      pos : "SUN_POS";
      plast : Date_And_Time;
   END_VAR
   VAR_TEMP
      tXCAL : "CALENDAR";
      tHOLIDAYS : Array[0..29] of "HOLIDAY_DATA";
      dtemp : DInt;
      tmp : Int;
   END_VAR
BEGIN


   #tXCAL := #XCAL;
   #tHOLIDAYS := #HOLIDAYS;

   IF #tXCAL.UTC T_COMP #last THEN
     (* run once per second *)
     (* update utc last calculated  *)
     #last := #tXCAL.UTC;
     #utod := T_CONV(#tXCAL.UTC);

     (* calculate ltc from utc *)
     #tXCAL.LDT := "UTC_TO_LTIME"(UTC:=#tXCAL.UTC, DST_ENABLE:=#tXCAL.DST_EN, TIME_ZONE_OFFSET:=#tXCAL.OFFSET);
     #tXCAL.LDATE := T_CONV(#tXCAL.LDT);
     #tXCAL.LTOD := T_CONV(#tXCAL.LDT);
     #dtemp := "DAY_OF_DATE"(#tXCAL.LDATE);
     #XCAL.NIGHT := #XCAL.LTOD < #XCAL.SUN_RISE OR #XCAL.LTOD > #XCAL.SUN_SET;

     (* run once per hour *)
     #tmp := "HOUR"(#tXCAL.LTOD);
     IF  #tmp <> #last_hour THEN
       #tXCAL.DST_ON := "DST"(#tXCAL.UTC) AND #tXCAL.DST_EN;
       #last_hour := #tmp;
     END_IF;

     (* run once per day *)
     IF #dtemp <> #last_day THEN
       #last_day := #dtemp;
       (* a new day has started, recalculate daily events *)
       #tXCAL.YEAR := "YEAR_OF_DATE"(#tXCAL.LDATE);
       #tXCAL.MONTH := "MONTH_OF_DATE"(#tXCAL.LDATE);
       #tXCAL.DAY := "DAY_OF_MONTH"(#tXCAL.LDATE);
       #tXCAL.WEEKDAY := "DAY_OF_WEEK"(#tXCAL.LDATE);
       #holy(DATE_IN := #tXCAL.LDATE, LANGU := #tXCAL.LANGUAGE, HOLIDAYS := #tHOLIDAYS);
       #tXCAL.HOLIDAY := #holy.Y;
       #tXCAL.HOLY_NAME BLKMOV #holy._NAME;
       #sun(LATITUDE := #tXCAL.LATITUDE, LONGITUDE := #tXCAL.LONGITUDE, UTC := T_CONV(#tXCAL.UTC), H := #H);
       #tXCAL.SUN_RISE := T_CONV(T_CONV(#sun.SUN_RISE) + #tXCAL.OFFSET * 60000 + SEL(G:=#tXCAL.DST_ON,IN0:=DINT#0,IN1:=3600000));
       #tXCAL.SUN_SET := T_CONV(T_CONV(#sun.SUN_SET) + #tXCAL.OFFSET * 60000 + SEL(G:=#tXCAL.DST_ON,IN0:=DINT#0,IN1:=3600000));
       #tXCAL.SUN_MIDDAY := T_CONV(T_CONV(#sun.MIDDAY) + #tXCAL.OFFSET * 60000 + SEL(G:=#tXCAL.DST_ON,IN0:=DINT#0,IN1:=3600000));
       #tXCAL.SUN_HEIGTH := #sun.SUN_DECLINATION;
       #tXCAL.WORK_WEEK := "WORK_WEEK"(#tXCAL.LDATE);
     END_IF;

     (* calculate the suns position every 10 seconds when SPE = TRUE *)
     IF #SPE AND #tXCAL.UTC T_DIFF #plast >= t#25s THEN
       #plast := #last;
       #pos(latitude := #tXCAL.LATITUDE, longitude := #tXCAL.LONGITUDE, utc := #tXCAL.UTC);
       #tXCAL.SUN_HOR := #pos."B";
       #tXCAL.SUN_VER := #pos.HR;
     END_IF;
   END_IF;

   #XCAL := #tXCAL;


   (* revision history

   hm 23. oct. 2008  rev 1.0
     original version

   hm  8. feb. 2009  rev 1.1
     night was calculated wrong
     added sun position data

   hm  10. mar. 2009 rev 1.2
     added work_week, sun_midday, sun_heigth
     sun_position will only be calculated evey 25 seconds
     dst will only become true when dst_en = true

   hm  23. jan 2010  rev 1.3
     sun_rise, sun_set and sun_midday are now calculated in local time

   hm  18. jan. 2011 rev 1.4
     added input holidays to specify local holidays
     changed call for function sun_time

   hm  2. feb. 2011  rev 1.5
     added input H to specify twilight

   hm  6. apr. 2011  rev 1.6
     night was calculated wrong
   *)
END_FUNCTION_BLOCK

FUNCTION_BLOCK "DCF77"   // FB27, SCL
TITLE = DCF77
{ S7_Optimized_Access := 'FALSE' }
AUTHOR : hugo
FAMILY : TIDT
NAME : DCF77
VERSION : 1.10
// this is a decoder for a DCF77 signal.
// the decoder decodes the DCF77 signal and checks for a valid Date_Time.
// since the dcf77 signal is only secured with a simple parity the decoder waits for two consecutive valid transmissions before it sets the output signals.
// given a valid reception by the receiver the decoder can take up to 3 minutes to start its clocks the first time.
// after a valid signal is detected the error output goes low and dignals a valid dcf signal from the receiver.
// a tp is only valid for one program cycle to allow for external rtc setting.
// after a valid signal is detected two independent internal clocks are started (RTC and RTC1), the seconds  of these clocks are generated by software since the dcf signal is only valid for minutes.
// rtc is always utc ( world time) and rtc1 can be set to any time zone by setting the time_zone_offset and enabling dst for automatic summertime.
// a sync output signals the the rtc and rtc1 are in sync with the dcf77 signal, if the dcf77 signal is lost for more then the sync time the sync output goes low
// but the rtc and rtc1 outputs keep running based on software timing until a valid dcf77 signal is received again and triggers the clock.
// in addition a millisecond output gives further resolutionof the clocks.
// a dst output shows if daylight saving time is enables and the weekday output shows which day of week currently is ( 1= monday ... 7= sunday).
// 
// uses: AD_DT_TM [FC1]
//       SB_DT_TM [FC35]
//       NE_DT [FC28]
//       GT_DT [FC14]
//       T_PLC_MS [FC64]
//       STIME [FB64],IDB_STIME [DB64]
//       EVEN [FC76]
//       DINT_DT [FC399]
//       D_TOD_DT [FC3] 
//       DT_DINT [FC400]
//       DT_DATE [FC6] 
//       DT_TOD [FC8] 
//       DAY_OF_WEEK [FC179]
//       DST [FC183]
//       YEAR_OF_DATE [FC219] 
//       SET_DT [FC214]
   VAR_INPUT
      REC : Bool;
      SET : Bool;
      SDT : Date_And_Time;
      DSI : Bool;
      SYNC_TIMEOUT : Time := T#2M;
      TIME_OFFSET : Int := 1;
      DST_EN : Bool := TRUE;
   END_VAR
   VAR_OUTPUT
      TP : Bool;
      DS : Bool;
      WDAY : Int;
      _WDAY AT WDAY : Array[0..15] of Bool;
      ERROR : Bool := TRUE;
      RTC : Date_And_Time;
      RTC1 : Date_And_Time;
      MSEC : Int;
      SYNC : Bool;
   END_VAR
   VAR
      MEZ : Date_And_Time;
      _MEZ AT MEZ : Struct
         Year : Byte;
         Month : Byte;
         Day : Byte;
         Hour : Byte;
         Minute : Byte;
         Second : Byte;
         ms : Byte;
         wday_ms : Byte;
      END_STRUCT;
      utc : Date_And_Time;
      state : Int;
      edge : Bool;
      tx : Time;
      ty : Time;
      last : Time;
      bits : Array[0..58] of Bool;
      cnt : Int;
      i : Int;
      old_time : Date_And_Time;
      minute : Byte;
      _minute AT minute : Array[0..7] of Bool;
      hour : Byte;
      _hour AT hour : Array[0..7] of Bool;
      day : Byte;
      _day AT day : Array[0..7] of Bool;
      month : Byte;
      _month AT month : Array[0..7] of Bool;
      year : Byte;
      _year AT year : Array[0..7] of Bool;
      last_sync : Time;
      t_1 : Time;
      tz : Time;
      init : Bool;
   END_VAR
   VAR_TEMP
      s7_wday : Int;
   END_VAR
BEGIN


     (* if tp was set it should only be active for 1 cycle *)
     #TP := FALSE;

     (* read system time *)
     #t_1 := T_CONV(DWORD_TO_DINT("T_PLC_MS"()));
     #tx := #t_1 - #last;

     IF #REC XOR #edge THEN
       #edge := #REC;
       IF NOT #REC AND #tx > t#1700ms AND #tx < t#2000ms THEN
         (* start condition reached *)
         #state := 0;
         #TP := NOT #ERROR;
       ELSIF NOT #REC AND #tx > t#700ms AND #tx < t#1000ms THEN
         (* second switch detected *)
         IF #state < 58 THEN #state := #state +1; ELSE #state := 0; END_IF;
       ELSIF #REC AND #tx  < t#120ms THEN
         (* bit 0 detected  *)
         #bits[#state] := 0;
       ELSIF #REC AND #tx > t#120ms AND #tx < t#250ms THEN
         (* bit 1 detected *)
         #bits[#state] := 1;
       ELSE
         (* error condition received signal is not valid *)
         #ERROR := TRUE;
         #state := 0;
       END_IF;
       #last := #last + #tx;
       IF #REC AND #state = 58 THEN
         #ERROR := FALSE;

         (* decode the bits and check for possible errors *)
         IF #bits[0] OR NOT (#bits[17] XOR #bits[18]) OR NOT #bits[20] THEN #ERROR := TRUE; END_IF;
         (* decode minute *)
         #minute := 0;
         #_minute[0] := #bits[21];
         #_minute[1] := #bits[22];
         #_minute[2] := #bits[23];
         #_minute[3] := #bits[24];
         #_minute[4] := #bits[25];
         #_minute[5] := #bits[26];
         #_minute[6] := #bits[27];
         IF BCD16_TO_INT(#minute) > 59 OR (#bits[21] XOR #bits[22] XOR #bits[23] XOR #bits[24] XOR #bits[25] XOR #bits[26] XOR #bits[27] XOR #bits[28]) THEN #ERROR := TRUE; END_IF;

         (* decode hour *)
         #hour := 0;
         #_hour[0] := #bits[29];
         #_hour[1] := #bits[30];
         #_hour[2] := #bits[31];
         #_hour[3] := #bits[32];
         #_hour[4] := #bits[33];
         #_hour[5] := #bits[34];
         IF BCD16_TO_INT(#hour) > 23 OR (#bits[29] XOR #bits[30] XOR #bits[31] XOR #bits[32] XOR #bits[33] XOR #bits[34] XOR #bits[35]) THEN #ERROR := TRUE; END_IF;

         (* decode day of month *)
         #day := 0;
         #_day[0] := #bits[36];
         #_day[1] := #bits[37];
         #_day[2] := #bits[38];
         #_day[3] := #bits[39];
         #_day[4] := #bits[40];
         #_day[5] := #bits[41];
         IF BCD16_TO_INT(#day) > 31 THEN #ERROR := TRUE; END_IF;

         (* decode day of week *)
         #WDAY := 0;
         #_WDAY[8] := #bits[42];
         #_WDAY[9] := #bits[43];
         #_WDAY[10] := #bits[44];
         IF #WDAY > 7 OR #WDAY < 1 THEN #ERROR := TRUE; END_IF;

         (* decode month *)
         #month := 0;
         #_month[0] := #bits[45];
         #_month[1] := #bits[46];
         #_month[2] := #bits[47];
         #_month[3] := #bits[48];
         #_month[4] := #bits[49];
         IF BCD16_TO_INT(#month) > 12 THEN #ERROR := TRUE; END_IF;

         (* decode year *)
         #year := 0;
         #_year[0] := #bits[50];
         #_year[1] := #bits[51];
         #_year[2] := #bits[52];
         #_year[3] := #bits[53];
         #_year[4] := #bits[54];
         #_year[5] := #bits[55];
         #_year[6] := #bits[56];
         #_year[7] := #bits[57];

         (* check parity for bits 36 to 58 *)
         #cnt := 0;
         FOR #i := 36 TO 58 DO IF #bits[#i] THEN #cnt := #cnt + 1; END_IF; END_FOR;
         IF NOT "EVEN"(#cnt) THEN #ERROR := TRUE; END_IF;

         (* time must be valid for two cycles to clear error flag *)
         IF NOT #ERROR THEN
           (* set outputs *)
           #old_time := #MEZ;
           //IF year >= 70 THEN year := year + 1900; ELSE year := year + 2000; END_IF;
           #_MEZ.Year := #year;
           #_MEZ.Month := #month;
           #_MEZ.Day := #day;
           #_MEZ.Hour := #hour;
           #_MEZ.Minute := #minute;
           #_MEZ.Second := 0;
           #_MEZ.ms := 0;

           //adaption S7 weekday Sunday is 1. 
           IF #WDAY < 7 THEN #s7_wday := #WDAY + 1; ELSE #s7_wday := 1; END_IF;
           #_MEZ.wday_ms := WORD_TO_BYTE(INT_TO_BCD16(#s7_wday));

           //mez := set_DT(year,month,day,hour,minute,0);
           #DS := #bits[17];
           IF #DS THEN
             #utc := "DINT_DT"("DT_DINT"(#MEZ) - 7200);
           ELSE
             #utc := "DINT_DT"("DT_DINT"(#MEZ) - 3600);
           END_IF;

           (* set trigger signal only if the receiver has received 2 successive minutes *)
           IF #MEZ T_COMP #old_time T_ADD t#1m THEN #ERROR := TRUE ; END_IF;
         END_IF;
       END_IF;
     END_IF;

     (* this portion implements a free running clock which is triggered by the dcf77 signal *)
     #tz := T_CONV(INT_TO_DINT(ABS(#TIME_OFFSET))* 3600000);

     IF NOT #init OR #SET THEN
       #init := TRUE;
       #utc := #SDT;
       #TP := TRUE;
       #DS := #DSI;
     END_IF;

     IF #TP THEN
       #RTC := #utc;
       IF #DS AND #DST_EN THEN
         IF #TIME_OFFSET < 0 THEN  #RTC1 := #RTC T_SUB #tz T_ADD t#1h; ELSE #RTC1 := #RTC T_ADD #tz T_ADD t#1h; END_IF;
       ELSE
         IF #TIME_OFFSET < 0 THEN #RTC1 := #RTC T_SUB #tz; ELSE #RTC1 := #RTC T_ADD #tz; END_IF;
       END_IF;
       #SYNC := TRUE;
       #last_sync := #last;
       #ty := #last;
     ELSIF #RTC T_COMP "DINT_DT"(0) AND #t_1 - #ty >= t#1s THEN
       #RTC := #RTC T_ADD t#1s;
       #RTC1 := #RTC1 T_ADD t#1s;
       #ty := #ty + t#1s;
       #SYNC := #ty - #last_sync < #SYNC_TIMEOUT AND #last_sync > T_CONV(0);
       #WDAY := "DAY_OF_WEEK"(T_CONV(#RTC1));
       #DS := #DST_EN AND "DST"(#utc);
     END_IF;
     #MSEC := DINT_TO_INT(T_CONV(#t_1 - #ty));



   (* decode information
   bits        content
   0           Bitwert immer 0
   1 bis 14    reserviert für Betriebsinformationen (nicht für DCF77-Nutzer bestimmt)
   15          Rufbit für Alarmierung der PTB-Mitarbeiter
               (bis Mai 2003: Bitwert = 0 falls normale Antenne in Verwendung; 1 = Backupantenne)
   16          Bitwert = 1 falls ein Wechsel von MEZ nach MESZ oder umgekehrt bevorsteht; Dauer der Anzeige: 1 Stunde
   17 + 18 gültige Zeit = MEZ, falls Bit 17=0 und Bit 18=1
               gültige Zeit = MESZ, falls Bit 17=1 und Bit 18=0
   19          Bitwert = 1 falls innerhalb den nächsten 59 Minuten eine Schaltsekunde angeordnet ist. Beim Einfügen einer Schaltsekunde wird anstelle der 59. die 60. Sekundenmarke weggelassen und in der 58. erfolgt ausnahmsweise ein Trägerabfall.
   20          Startbit für Zeitinformation (immer 1)
   21 - 27     1, 2, 4, 8, 10, 20, 40 Minuten (bitweise Addition)
   28          Prüfbit (gerade Parität) für die Bits 21-27
   29 - 34     1, 2, 4, 8, 10, 20 Stunden (bitweise Addition)
   35          Prüfbit (gerade Parität) für die Bits 29-34
   36 - 41     Tagesnummer im aktuellen Monat: 1, 2, 4, 8, 10, 20 (bitweise Addition)
   42 - 44     Tagesnummer in der aktuellen Woche: 1, 2, 4 (bitweise Addition)
   45 - 49     Monatsnummer: 1, 2, 4, 8, 10 (bitweise Addition)
   50 - 57     Jahr (zweistellig): 1, 2, 4, 8, 10, 20, 40, 80 (bitweise Addition)
   58          Prüfbit (gerade Parität) füR die Bits 36-57

   *)
   (* revision history

   hm 2.feb 2007       rev 1.1
       change wday and dst outputs when there is no dcf reception

   hm  26.feb 2007     rev 1.2
       changed statements where t#1h would be substracted from DT.
       under certain conditions the compiler would crash translating this statement

   hm  17. sep 2007    rev 1.3
       replaced time() with T_PLC_MS() for compatibility reasons